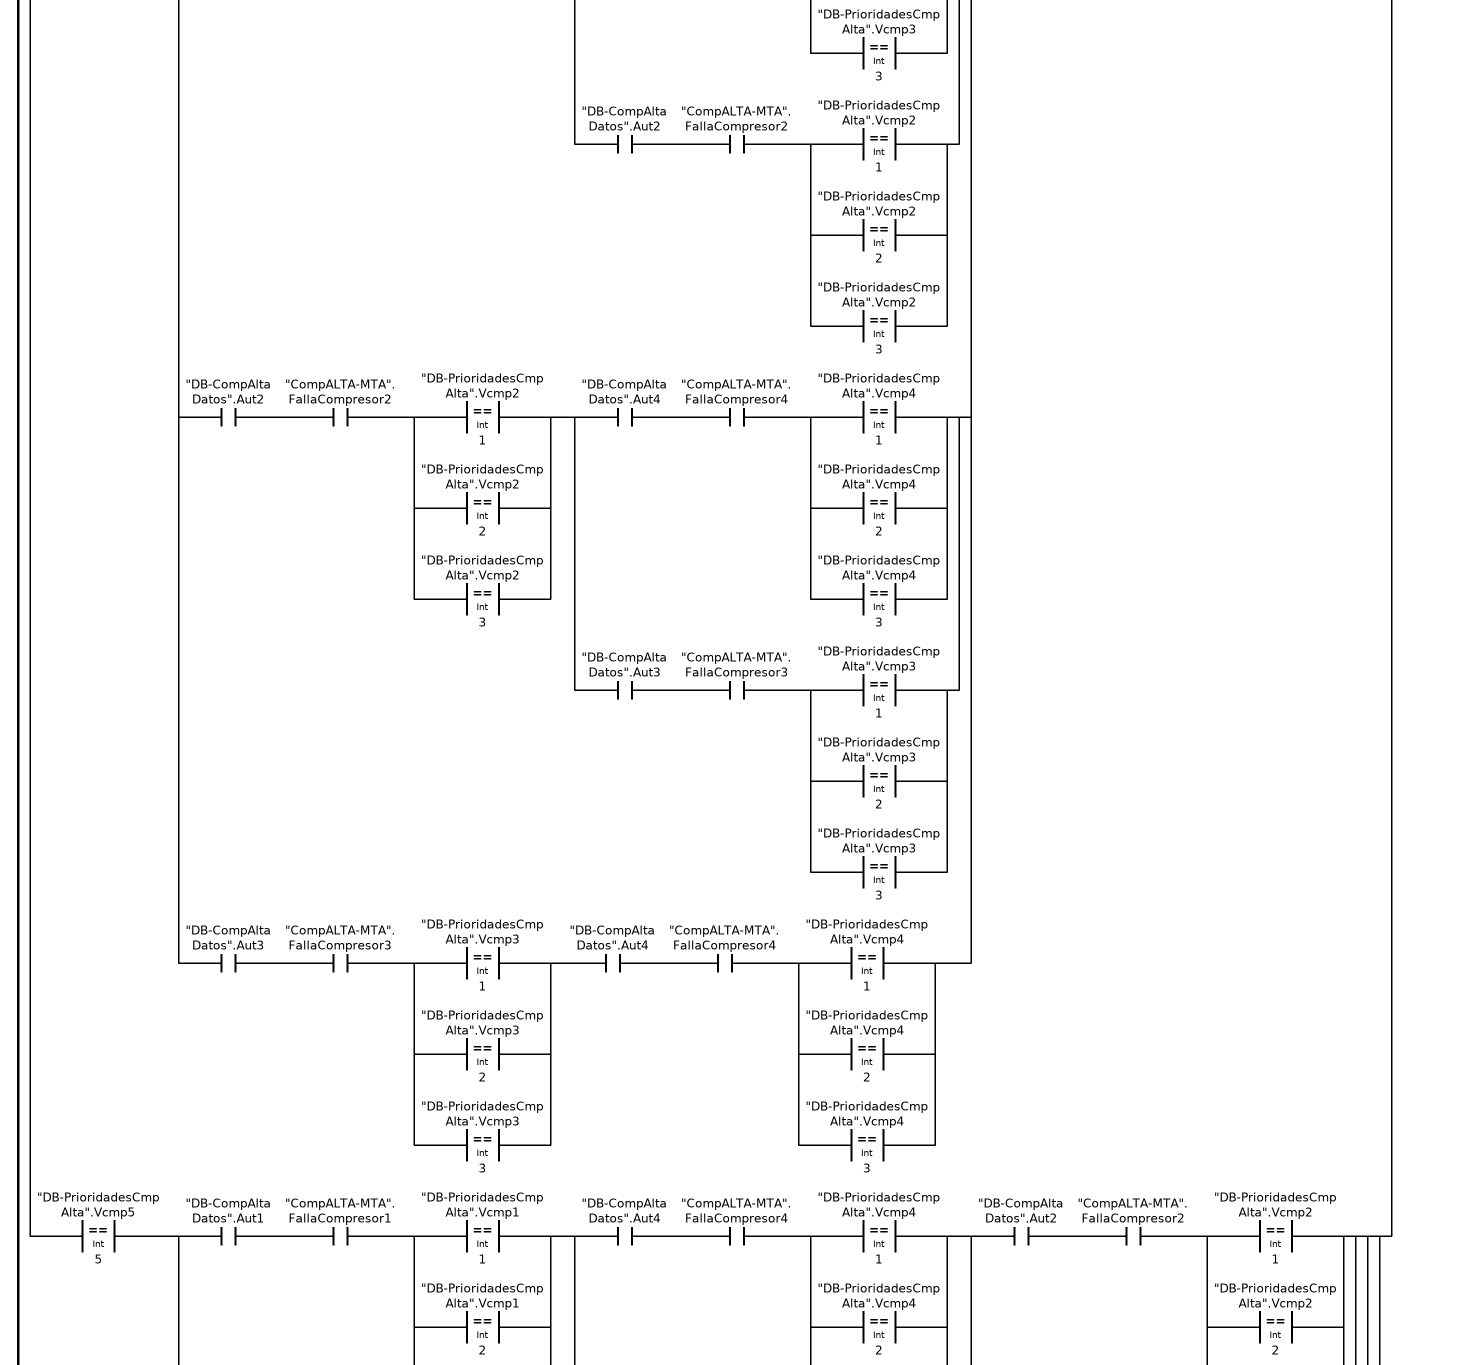
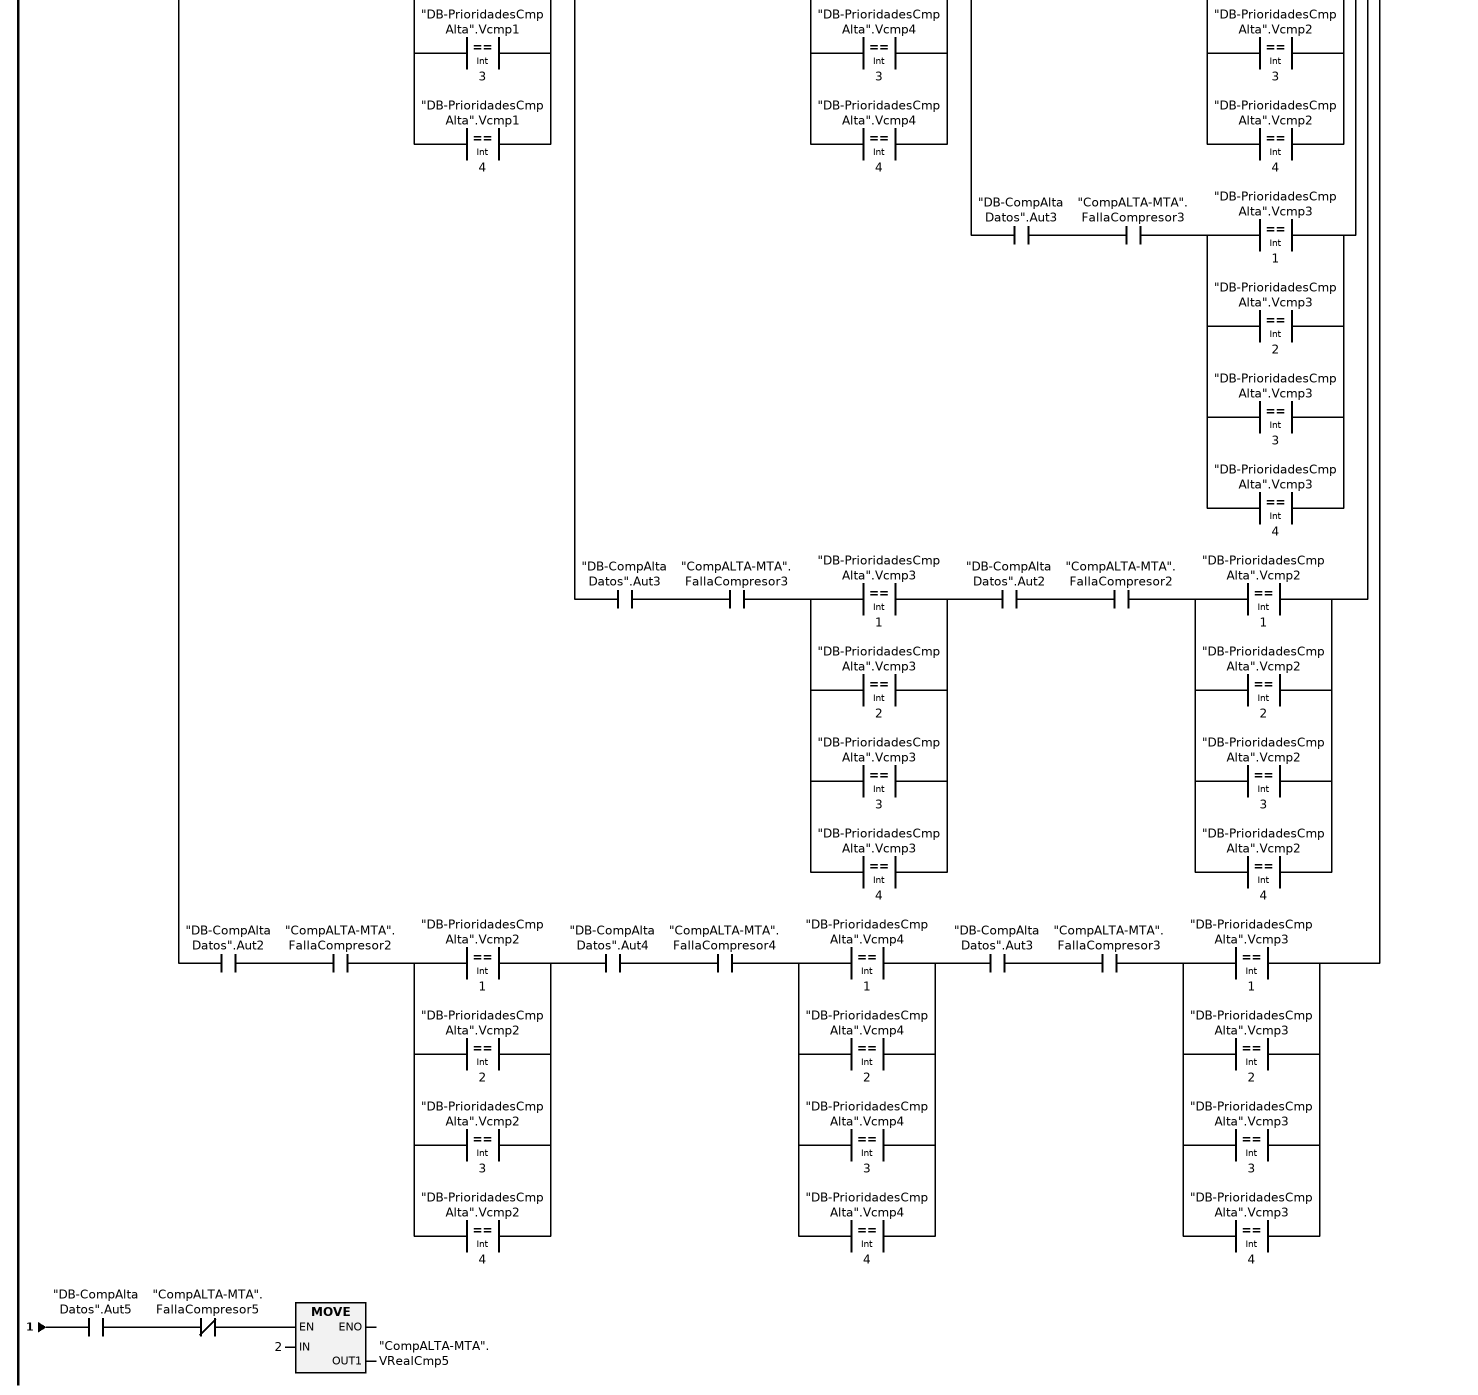
   IF (("DB-PrioridadesCmpAlta".Vcmp5 = 2) OR (("DB-PrioridadesCmpAlta".Vcmp5 = 3) AND (("DB-CompAltaDatos".Aut1 AND "CompALTA-MTA".FallaCompresor1 AND (("DB-PrioridadesCmpAlta".Vcmp1 = 2) OR ("DB-PrioridadesCmpAlta".Vcmp1 = 1))) OR ("DB-CompAltaDatos".Aut2 AND "CompALTA-MTA".FallaCompresor2 AND (("DB-PrioridadesCmpAlta".Vcmp2 = 2) OR ("DB-PrioridadesCmpAlta".Vcmp2 = 1))) OR ("DB-CompAltaDatos".Aut3 AND "CompALTA-MTA".FallaCompresor3 AND (("DB-PrioridadesCmpAlta".Vcmp3 = 2) OR ("DB-PrioridadesCmpAlta".Vcmp3 = 1))) OR ("DB-CompAltaDatos".Aut4 AND "CompALTA-MTA".FallaCompresor4 AND (("DB-PrioridadesCmpAlta".Vcmp4 = 2) OR ("DB-PrioridadesCmpAlta".Vcmp4 = 1))))) OR (("DB-PrioridadesCmpAlta".Vcmp5 = 4) AND (("DB-CompAltaDatos".Aut1 AND "CompALTA-MTA".FallaCompresor1 AND (("DB-PrioridadesCmpAlta".Vcmp1 = 1) OR ("DB-PrioridadesCmpAlta".Vcmp1 = 2) OR ("DB-PrioridadesCmpAlta".Vcmp1 = 3)) AND (("DB-CompAltaDatos".Aut4 AND "CompALTA-MTA".FallaCompresor4 AND (("DB-PrioridadesCmpAlta".Vcmp4 = 1) OR ("DB-PrioridadesCmpAlta".Vcmp4 = 2) OR ("DB-PrioridadesCmpAlta".Vcmp4 = 3))) OR ("DB-CompAltaDatos".Aut3 AND "CompALTA-MTA".FallaCompresor3 AND (("DB-PrioridadesCmpAlta".Vcmp3 = 1) OR ("DB-PrioridadesCmpAlta".Vcmp3 = 2) OR ("DB-PrioridadesCmpAlta".Vcmp3 = 3))) OR ("DB-CompAltaDatos".Aut2 AND "CompALTA-MTA".FallaCompresor2 AND (("DB-PrioridadesCmpAlta".Vcmp2 = 1) OR ("DB-PrioridadesCmpAlta".Vcmp2 = 2) OR ("DB-PrioridadesCmpAlta".Vcmp2 = 3))))) OR ("DB-CompAltaDatos".Aut2 AND "CompALTA-MTA".FallaCompresor2 AND (("DB-PrioridadesCmpAlta".Vcmp2 = 1) OR ("DB-PrioridadesCmpAlta".Vcmp2 = 2) OR ("DB-PrioridadesCmpAlta".Vcmp2 = 3)) AND (("DB-CompAltaDatos".Aut4 AND "CompALTA-MTA".FallaCompresor4 AND (("DB-PrioridadesCmpAlta".Vcmp4 = 1) OR ("DB-PrioridadesCmpAlta".Vcmp4 = 2) OR ("DB-PrioridadesCmpAlta".Vcmp4 = 3))) OR ("DB-CompAltaDatos".Aut3 AND "CompALTA-MTA".FallaCompresor3 AND (("DB-PrioridadesCmpAlta".Vcmp3 = 1) OR ("DB-PrioridadesCmpAlta".Vcmp3 = 2) OR ("DB-PrioridadesCmpAlta".Vcmp3 = 3))))) OR ("DB-CompAltaDatos".Aut3 AND "CompALTA-MTA".FallaCompresor3 AND (("DB-PrioridadesCmpAlta".Vcmp3 = 1) OR ("DB-PrioridadesCmpAlta".Vcmp3 = 2) OR ("DB-PrioridadesCmpAlta".Vcmp3 = 3)) AND "DB-CompAltaDatos".Aut4 AND "CompALTA-MTA".FallaCompresor4 AND (("DB-PrioridadesCmpAlta".Vcmp4 = 1) OR ("DB-PrioridadesCmpAlta".Vcmp4 = 2) OR ("DB-PrioridadesCmpAlta".Vcmp4 = 3))))) OR (("DB-PrioridadesCmpAlta".Vcmp5 = 5) AND (("DB-CompAltaDatos".Aut1 AND "CompALTA-MTA".FallaCompresor1 AND (("DB-PrioridadesCmpAlta".Vcmp1 = 1) OR ("DB-PrioridadesCmpAlta".Vcmp1 = 2) OR ("DB-PrioridadesCmpAlta".Vcmp1 = 3) OR ("DB-PrioridadesCmpAlta".Vcmp1 = 4)) AND (("DB-CompAltaDatos".Aut4 AND "CompALTA-MTA".FallaCompresor4 AND (("DB-PrioridadesCmpAlta".Vcmp4 = 1) OR ("DB-PrioridadesCmpAlta".Vcmp4 = 2) OR ("DB-PrioridadesCmpAlta".Vcmp4 = 3) OR ("DB-PrioridadesCmpAlta".Vcmp4 = 4)) AND (("DB-CompAltaDatos".Aut2 AND "CompALTA-MTA".FallaCompresor2 AND (("DB-PrioridadesCmpAlta".Vcmp2 = 1) OR ("DB-PrioridadesCmpAlta".Vcmp2 = 2) OR ("DB-PrioridadesCmpAlta".Vcmp2 = 3) OR ("DB-PrioridadesCmpAlta".Vcmp2 = 4))) OR ("DB-CompAltaDatos".Aut3 AND "CompALTA-MTA".FallaCompresor3 AND (("DB-PrioridadesCmpAlta".Vcmp3 = 1) OR ("DB-PrioridadesCmpAlta".Vcmp3 = 2) OR ("DB-PrioridadesCmpAlta".Vcmp3 = 3) OR ("DB-PrioridadesCmpAlta".Vcmp3 = 4))))) OR ("DB-CompAltaDatos".Aut3 AND "CompALTA-MTA".FallaCompresor3 AND (("DB-PrioridadesCmpAlta".Vcmp3 = 1) OR ("DB-PrioridadesCmpAlta".Vcmp3 = 2) OR ("DB-PrioridadesCmpAlta".Vcmp3 = 3) OR ("DB-PrioridadesCmpAlta".Vcmp3 = 4)) AND "DB-CompAltaDatos".Aut2 AND "CompALTA-MTA".FallaCompresor2 AND (("DB-PrioridadesCmpAlta".Vcmp2 = 1) OR ("DB-PrioridadesCmpAlta".Vcmp2 = 2) OR ("DB-PrioridadesCmpAlta".Vcmp2 = 3) OR ("DB-PrioridadesCmpAlta".Vcmp2 = 4))))) OR ("DB-CompAltaDatos".Aut2 AND "CompALTA-MTA".FallaCompresor2 AND (("DB-PrioridadesCmpAlta".Vcmp2 = 1) OR ("DB-PrioridadesCmpAlta".Vcmp2 = 2) OR ("DB-PrioridadesCmpAlta".Vcmp2 = 3) OR ("DB-PrioridadesCmpAlta".Vcmp2 = 4)) AND "DB-CompAltaDatos".Aut4 AND "CompALTA-MTA".FallaCompresor4 AND (("DB-PrioridadesCmpAlta".Vcmp4 = 1) OR ("DB-PrioridadesCmpAlta".Vcmp4 = 2) OR ("DB-PrioridadesCmpAlta".Vcmp4 = 3) OR ("DB-PrioridadesCmpAlta".Vcmp4 = 4)) AND "DB-CompAltaDatos".Aut3 AND "CompALTA-MTA".FallaCompresor3 AND (("DB-PrioridadesCmpAlta".Vcmp3 = 1) OR ("DB-PrioridadesCmpAlta".Vcmp3 = 2) OR ("DB-PrioridadesCmpAlta".Vcmp3 = 3) OR ("DB-PrioridadesCmpAlta".Vcmp3 = 4)))))) AND "DB-CompAltaDatos".Aut5 AND NOT "CompALTA-MTA".FallaCompresor5 THEN
       "CompALTA-MTA".VRealCmp5 := 2;
   END_IF;
END_REGION

REGION Network 33
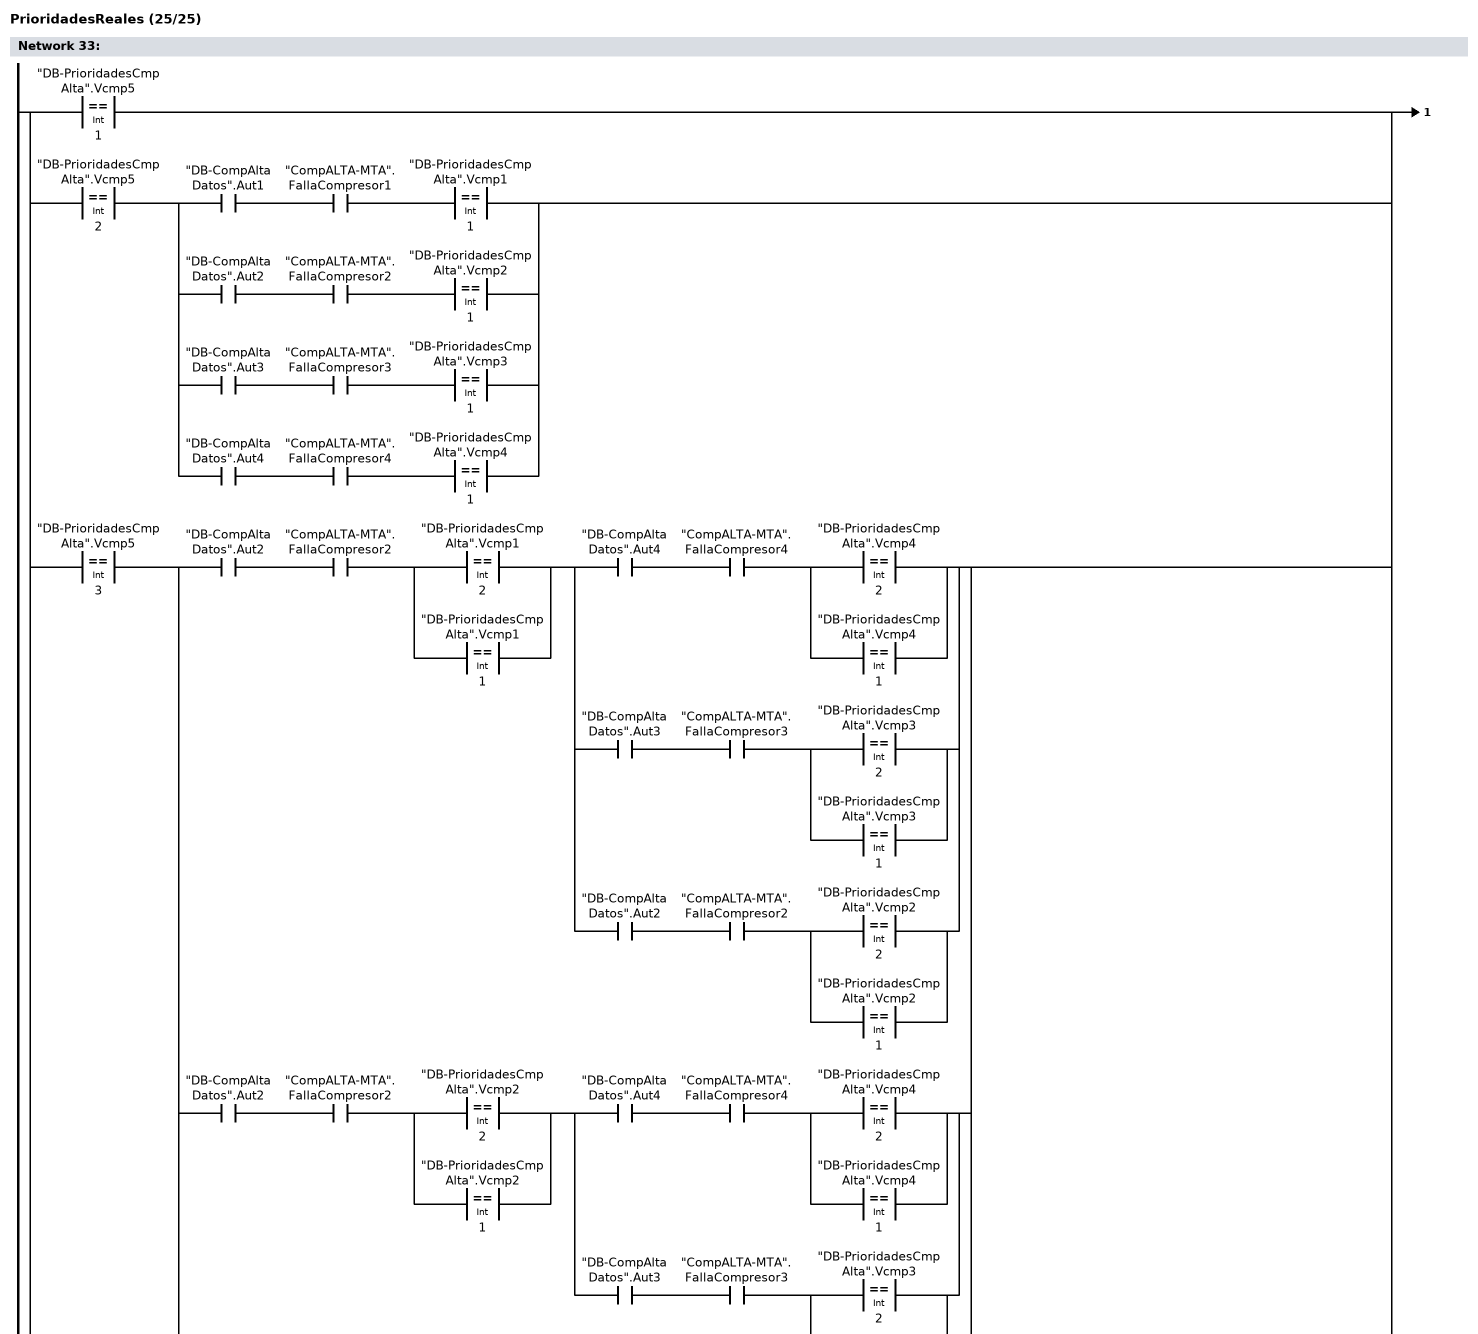
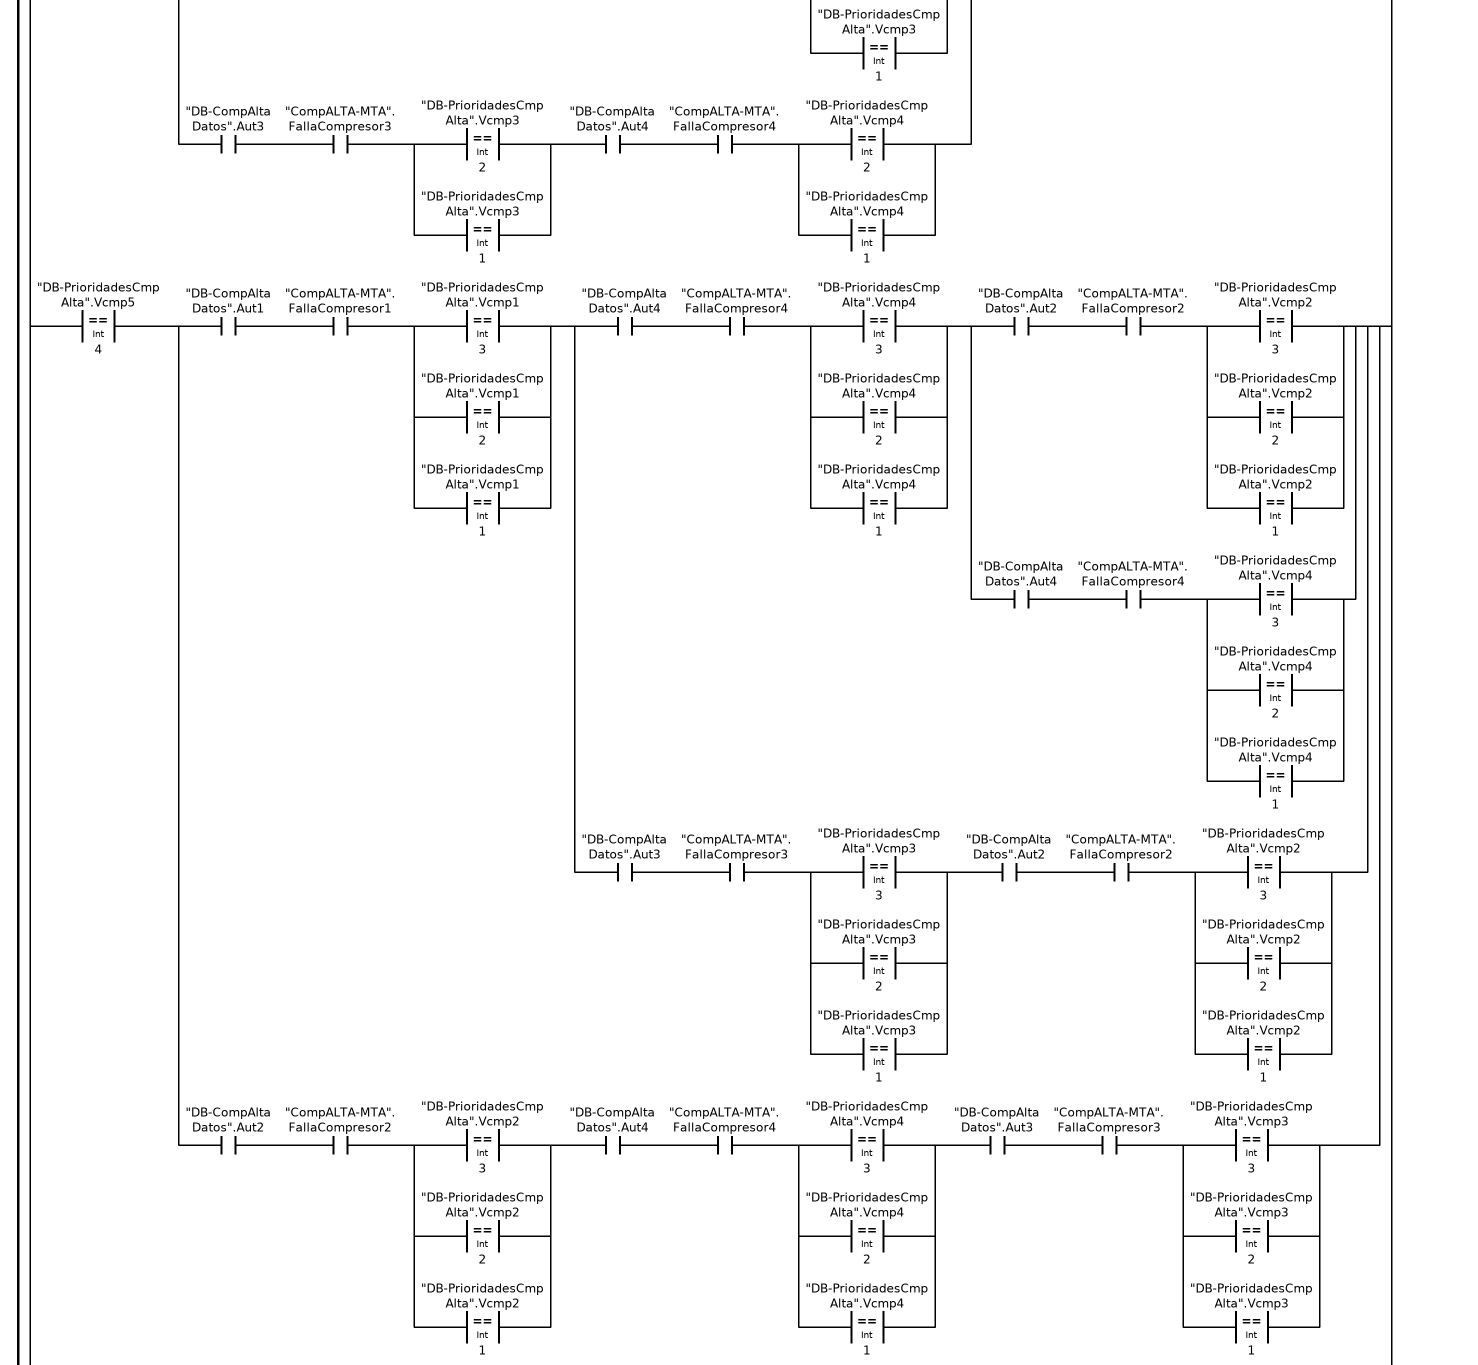
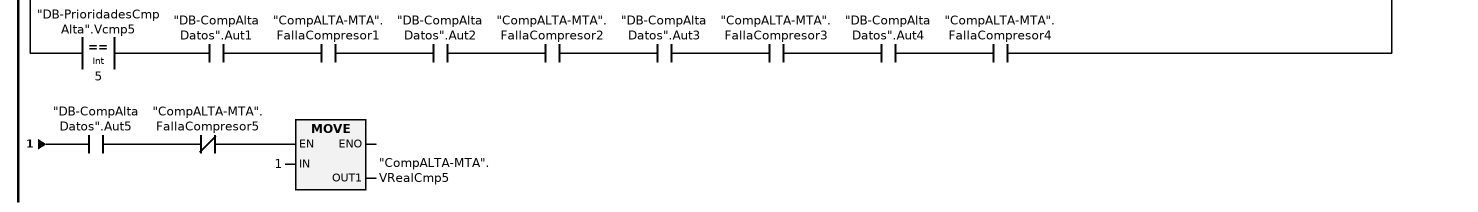
   IF (("DB-PrioridadesCmpAlta".Vcmp5 = 1) OR (("DB-PrioridadesCmpAlta".Vcmp5 = 2) AND (("DB-CompAltaDatos".Aut1 AND "CompALTA-MTA".FallaCompresor1 AND ("DB-PrioridadesCmpAlta".Vcmp1 = 1)) OR ("DB-CompAltaDatos".Aut2 AND "CompALTA-MTA".FallaCompresor2 AND ("DB-PrioridadesCmpAlta".Vcmp2 = 1)) OR ("DB-CompAltaDatos".Aut3 AND "CompALTA-MTA".FallaCompresor3 AND ("DB-PrioridadesCmpAlta".Vcmp3 = 1)) OR ("DB-CompAltaDatos".Aut4 AND "CompALTA-MTA".FallaCompresor4 AND ("DB-PrioridadesCmpAlta".Vcmp4 = 1)))) OR (("DB-PrioridadesCmpAlta".Vcmp5 = 3) AND (("DB-CompAltaDatos".Aut2 AND "CompALTA-MTA".FallaCompresor2 AND (("DB-PrioridadesCmpAlta".Vcmp1 = 2) OR ("DB-PrioridadesCmpAlta".Vcmp1 = 1)) AND (("DB-CompAltaDatos".Aut4 AND "CompALTA-MTA".FallaCompresor4 AND (("DB-PrioridadesCmpAlta".Vcmp4 = 2) OR ("DB-PrioridadesCmpAlta".Vcmp4 = 1))) OR ("DB-CompAltaDatos".Aut3 AND "CompALTA-MTA".FallaCompresor3 AND (("DB-PrioridadesCmpAlta".Vcmp3 = 2) OR ("DB-PrioridadesCmpAlta".Vcmp3 = 1))) OR ("DB-CompAltaDatos".Aut2 AND "CompALTA-MTA".FallaCompresor2 AND (("DB-PrioridadesCmpAlta".Vcmp2 = 2) OR ("DB-PrioridadesCmpAlta".Vcmp2 = 1))))) OR ("DB-CompAltaDatos".Aut2 AND "CompALTA-MTA".FallaCompresor2 AND (("DB-PrioridadesCmpAlta".Vcmp2 = 2) OR ("DB-PrioridadesCmpAlta".Vcmp2 = 1)) AND (("DB-CompAltaDatos".Aut4 AND "CompALTA-MTA".FallaCompresor4 AND (("DB-PrioridadesCmpAlta".Vcmp4 = 2) OR ("DB-PrioridadesCmpAlta".Vcmp4 = 1))) OR ("DB-CompAltaDatos".Aut3 AND "CompALTA-MTA".FallaCompresor3 AND (("DB-PrioridadesCmpAlta".Vcmp3 = 2) OR ("DB-PrioridadesCmpAlta".Vcmp3 = 1))))) OR ("DB-CompAltaDatos".Aut3 AND "CompALTA-MTA".FallaCompresor3 AND (("DB-PrioridadesCmpAlta".Vcmp3 = 2) OR ("DB-PrioridadesCmpAlta".Vcmp3 = 1)) AND "DB-CompAltaDatos".Aut4 AND "CompALTA-MTA".FallaCompresor4 AND (("DB-PrioridadesCmpAlta".Vcmp4 = 2) OR ("DB-PrioridadesCmpAlta".Vcmp4 = 1))))) OR (("DB-PrioridadesCmpAlta".Vcmp5 = 4) AND (("DB-CompAltaDatos".Aut1 AND "CompALTA-MTA".FallaCompresor1 AND (("DB-PrioridadesCmpAlta".Vcmp1 = 3) OR ("DB-PrioridadesCmpAlta".Vcmp1 = 2) OR ("DB-PrioridadesCmpAlta".Vcmp1 = 1)) AND (("DB-CompAltaDatos".Aut4 AND "CompALTA-MTA".FallaCompresor4 AND (("DB-PrioridadesCmpAlta".Vcmp4 = 3) OR ("DB-PrioridadesCmpAlta".Vcmp4 = 2) OR ("DB-PrioridadesCmpAlta".Vcmp4 = 1)) AND (("DB-CompAltaDatos".Aut2 AND "CompALTA-MTA".FallaCompresor2 AND (("DB-PrioridadesCmpAlta".Vcmp2 = 3) OR ("DB-PrioridadesCmpAlta".Vcmp2 = 2) OR ("DB-PrioridadesCmpAlta".Vcmp2 = 1))) OR ("DB-CompAltaDatos".Aut4 AND "CompALTA-MTA".FallaCompresor4 AND (("DB-PrioridadesCmpAlta".Vcmp4 = 3) OR ("DB-PrioridadesCmpAlta".Vcmp4 = 2) OR ("DB-PrioridadesCmpAlta".Vcmp4 = 1))))) OR ("DB-CompAltaDatos".Aut3 AND "CompALTA-MTA".FallaCompresor3 AND (("DB-PrioridadesCmpAlta".Vcmp3 = 3) OR ("DB-PrioridadesCmpAlta".Vcmp3 = 2) OR ("DB-PrioridadesCmpAlta".Vcmp3 = 1)) AND "DB-CompAltaDatos".Aut2 AND "CompALTA-MTA".FallaCompresor2 AND (("DB-PrioridadesCmpAlta".Vcmp2 = 3) OR ("DB-PrioridadesCmpAlta".Vcmp2 = 2) OR ("DB-PrioridadesCmpAlta".Vcmp2 = 1))))) OR ("DB-CompAltaDatos".Aut2 AND "CompALTA-MTA".FallaCompresor2 AND (("DB-PrioridadesCmpAlta".Vcmp2 = 3) OR ("DB-PrioridadesCmpAlta".Vcmp2 = 2) OR ("DB-PrioridadesCmpAlta".Vcmp2 = 1)) AND "DB-CompAltaDatos".Aut4 AND "CompALTA-MTA".FallaCompresor4 AND (("DB-PrioridadesCmpAlta".Vcmp4 = 3) OR ("DB-PrioridadesCmpAlta".Vcmp4 = 2) OR ("DB-PrioridadesCmpAlta".Vcmp4 = 1)) AND "DB-CompAltaDatos".Aut3 AND "CompALTA-MTA".FallaCompresor3 AND (("DB-PrioridadesCmpAlta".Vcmp3 = 3) OR ("DB-PrioridadesCmpAlta".Vcmp3 = 2) OR ("DB-PrioridadesCmpAlta".Vcmp3 = 1))))) OR (("DB-PrioridadesCmpAlta".Vcmp5 = 5) AND "DB-CompAltaDatos".Aut1 AND "CompALTA-MTA".FallaCompresor1 AND "DB-CompAltaDatos".Aut2 AND "CompALTA-MTA".FallaCompresor2 AND "DB-CompAltaDatos".Aut3 AND "CompALTA-MTA".FallaCompresor3 AND "DB-CompAltaDatos".Aut4 AND "CompALTA-MTA".FallaCompresor4)) AND "DB-CompAltaDatos".Aut5 AND NOT "CompALTA-MTA".FallaCompresor5 THEN
       "CompALTA-MTA".VRealCmp5 := 1;
   END_IF;
END_REGION
END_FUNCTION

FUNCTION "FlancosCmpAlta" : Void   // FC45, LAD
{ S7_Optimized_Access := 'FALSE' }
VERSION : 0.1
   VAR_TEMP   // added for the SCL form of the ladder/FBD networks
      _w1 : Bool;
      _w2 : Bool;
      _w3 : Bool;
      _w4 : Bool;
      _w5 : Bool;
      _w6 : Bool;
      _w7 : Bool;
      _s5time1 : S5Time;
   END_VAR
BEGIN

REGION Network 1
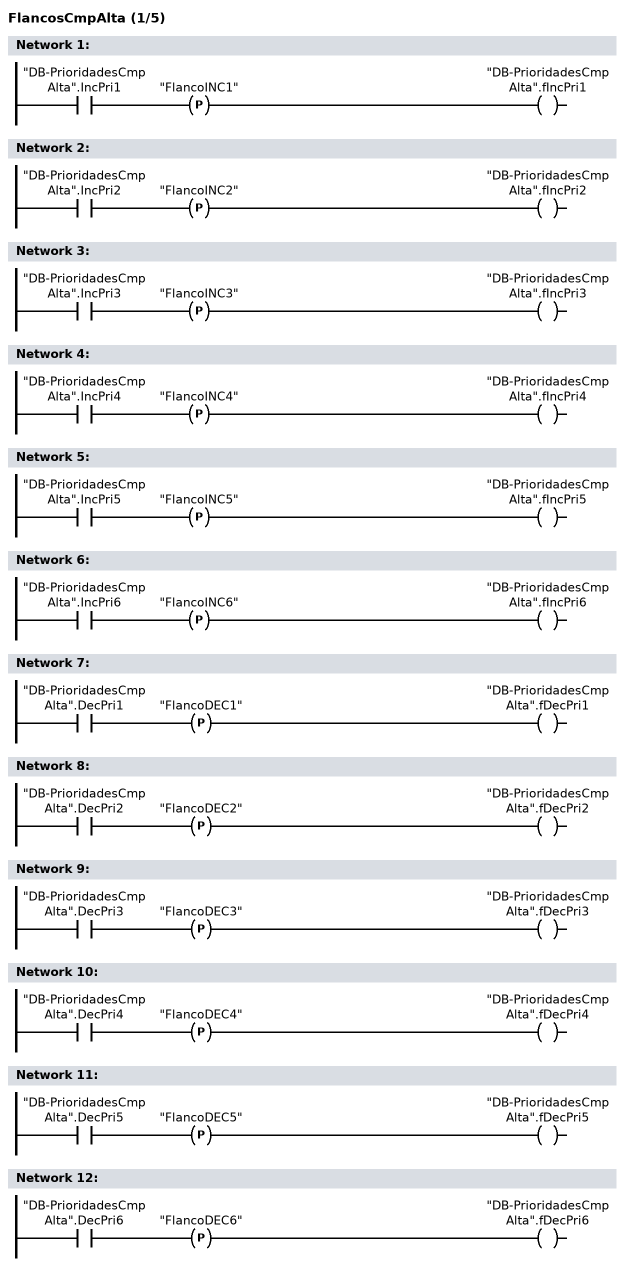
   RUNG wire#powerrail
      Contact( "DB-PrioridadesCmpAlta".IncPri1 )
      P_Trig( "FlancoINC1" )
      Coil( "DB-PrioridadesCmpAlta".fIncPri1 )
   END_RUNG
   // the same network as SCL:
   #_w1 := "DB-PrioridadesCmpAlta".IncPri1 AND NOT "FlancoINC1";   // rising edge
   "FlancoINC1" := "DB-PrioridadesCmpAlta".IncPri1;
   "DB-PrioridadesCmpAlta".fIncPri1 := #_w1;
END_REGION

REGION Network 2
   RUNG wire#powerrail
      Contact( "DB-PrioridadesCmpAlta".IncPri2 )
      P_Trig( "FlancoINC2" )
      Coil( "DB-PrioridadesCmpAlta".fIncPri2 )
   END_RUNG
   // the same network as SCL:
   #_w1 := "DB-PrioridadesCmpAlta".IncPri2 AND NOT "FlancoINC2";   // rising edge
   "FlancoINC2" := "DB-PrioridadesCmpAlta".IncPri2;
   "DB-PrioridadesCmpAlta".fIncPri2 := #_w1;
END_REGION

REGION Network 3
   RUNG wire#powerrail
      Contact( "DB-PrioridadesCmpAlta".IncPri3 )
      P_Trig( "FlancoINC3" )
      Coil( "DB-PrioridadesCmpAlta".fIncPri3 )
   END_RUNG
   // the same network as SCL:
   #_w1 := "DB-PrioridadesCmpAlta".IncPri3 AND NOT "FlancoINC3";   // rising edge
   "FlancoINC3" := "DB-PrioridadesCmpAlta".IncPri3;
   "DB-PrioridadesCmpAlta".fIncPri3 := #_w1;
END_REGION

REGION Network 4
   RUNG wire#powerrail
      Contact( "DB-PrioridadesCmpAlta".IncPri4 )
      P_Trig( "FlancoINC4" )
      Coil( "DB-PrioridadesCmpAlta".fIncPri4 )
   END_RUNG
   // the same network as SCL:
   #_w1 := "DB-PrioridadesCmpAlta".IncPri4 AND NOT "FlancoINC4";   // rising edge
   "FlancoINC4" := "DB-PrioridadesCmpAlta".IncPri4;
   "DB-PrioridadesCmpAlta".fIncPri4 := #_w1;
END_REGION

REGION Network 5
   RUNG wire#powerrail
      Contact( "DB-PrioridadesCmpAlta".IncPri5 )
      P_Trig( "FlancoINC5" )
      Coil( "DB-PrioridadesCmpAlta".fIncPri5 )
   END_RUNG
   // the same network as SCL:
   #_w1 := "DB-PrioridadesCmpAlta".IncPri5 AND NOT "FlancoINC5";   // rising edge
   "FlancoINC5" := "DB-PrioridadesCmpAlta".IncPri5;
   "DB-PrioridadesCmpAlta".fIncPri5 := #_w1;
END_REGION

REGION Network 6
   RUNG wire#powerrail
      Contact( "DB-PrioridadesCmpAlta".IncPri6 )
      P_Trig( "FlancoINC6" )
      Coil( "DB-PrioridadesCmpAlta".fIncPri6 )
   END_RUNG
   // the same network as SCL:
   #_w1 := "DB-PrioridadesCmpAlta".IncPri6 AND NOT "FlancoINC6";   // rising edge
   "FlancoINC6" := "DB-PrioridadesCmpAlta".IncPri6;
   "DB-PrioridadesCmpAlta".fIncPri6 := #_w1;
END_REGION

REGION Network 7
   RUNG wire#powerrail
      Contact( "DB-PrioridadesCmpAlta".DecPri1 )
      P_Trig( "FlancoDEC1" )
      Coil( "DB-PrioridadesCmpAlta".fDecPri1 )
   END_RUNG
   // the same network as SCL:
   #_w1 := "DB-PrioridadesCmpAlta".DecPri1 AND NOT "FlancoDEC1";   // rising edge
   "FlancoDEC1" := "DB-PrioridadesCmpAlta".DecPri1;
   "DB-PrioridadesCmpAlta".fDecPri1 := #_w1;
END_REGION

REGION Network 8
   RUNG wire#powerrail
      Contact( "DB-PrioridadesCmpAlta".DecPri2 )
      P_Trig( "FlancoDEC2" )
      Coil( "DB-PrioridadesCmpAlta".fDecPri2 )
   END_RUNG
   // the same network as SCL:
   #_w1 := "DB-PrioridadesCmpAlta".DecPri2 AND NOT "FlancoDEC2";   // rising edge
   "FlancoDEC2" := "DB-PrioridadesCmpAlta".DecPri2;
   "DB-PrioridadesCmpAlta".fDecPri2 := #_w1;
END_REGION

REGION Network 9
   RUNG wire#powerrail
      Contact( "DB-PrioridadesCmpAlta".DecPri3 )
      P_Trig( "FlancoDEC3" )
      Coil( "DB-PrioridadesCmpAlta".fDecPri3 )
   END_RUNG
   // the same network as SCL:
   #_w1 := "DB-PrioridadesCmpAlta".DecPri3 AND NOT "FlancoDEC3";   // rising edge
   "FlancoDEC3" := "DB-PrioridadesCmpAlta".DecPri3;
   "DB-PrioridadesCmpAlta".fDecPri3 := #_w1;
END_REGION

REGION Network 10
   RUNG wire#powerrail
      Contact( "DB-PrioridadesCmpAlta".DecPri4 )
      P_Trig( "FlancoDEC4" )
      Coil( "DB-PrioridadesCmpAlta".fDecPri4 )
   END_RUNG
   // the same network as SCL:
   #_w1 := "DB-PrioridadesCmpAlta".DecPri4 AND NOT "FlancoDEC4";   // rising edge
   "FlancoDEC4" := "DB-PrioridadesCmpAlta".DecPri4;
   "DB-PrioridadesCmpAlta".fDecPri4 := #_w1;
END_REGION

REGION Network 11
   RUNG wire#powerrail
      Contact( "DB-PrioridadesCmpAlta".DecPri5 )
      P_Trig( "FlancoDEC5" )
      Coil( "DB-PrioridadesCmpAlta".fDecPri5 )
   END_RUNG
   // the same network as SCL:
   #_w1 := "DB-PrioridadesCmpAlta".DecPri5 AND NOT "FlancoDEC5";   // rising edge
   "FlancoDEC5" := "DB-PrioridadesCmpAlta".DecPri5;
   "DB-PrioridadesCmpAlta".fDecPri5 := #_w1;
END_REGION

REGION Network 12
   RUNG wire#powerrail
      Contact( "DB-PrioridadesCmpAlta".DecPri6 )
      P_Trig( "FlancoDEC6" )
      Coil( "DB-PrioridadesCmpAlta".fDecPri6 )
   END_RUNG
   // the same network as SCL:
   #_w1 := "DB-PrioridadesCmpAlta".DecPri6 AND NOT "FlancoDEC6";   // rising edge
   "FlancoDEC6" := "DB-PrioridadesCmpAlta".DecPri6;
   "DB-PrioridadesCmpAlta".fDecPri6 := #_w1;
END_REGION

REGION Network 13
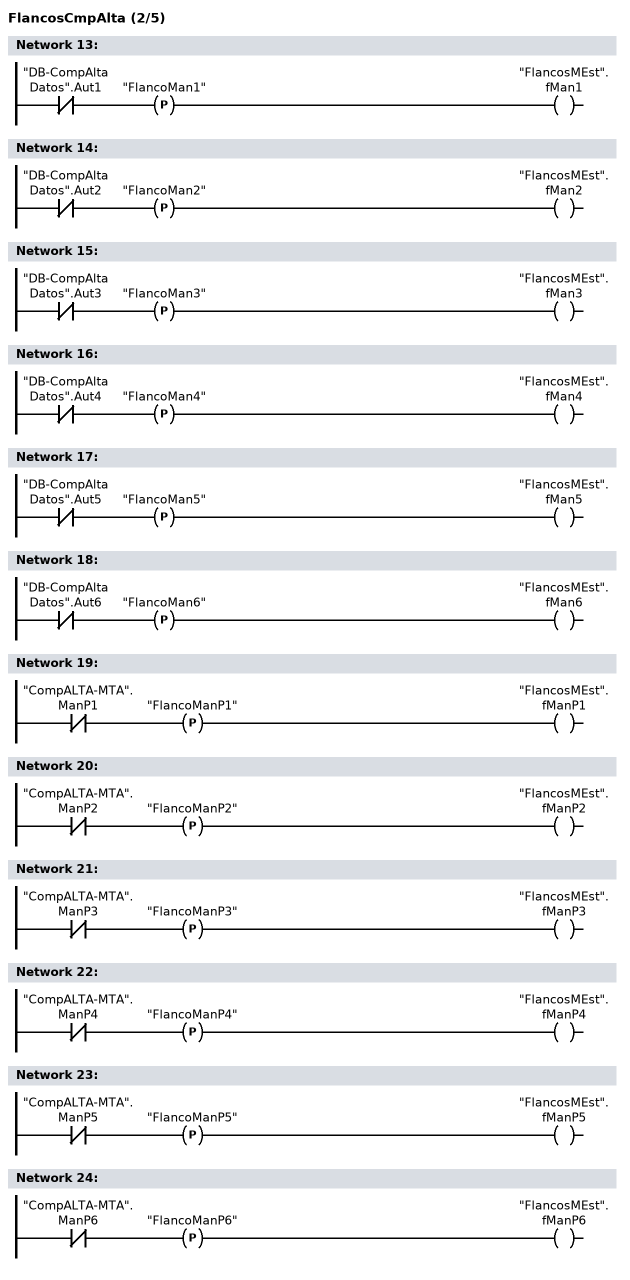
   RUNG wire#powerrail
      I_Contact( "DB-CompAltaDatos".Aut1 )
      P_Trig( "FlancoMan1" )
      Coil( "FlancosMEst".fMan1 )
   END_RUNG
   // the same network as SCL:
   #_w1 := NOT "DB-CompAltaDatos".Aut1 AND NOT "FlancoMan1";   // rising edge
   "FlancoMan1" := NOT "DB-CompAltaDatos".Aut1;
   "FlancosMEst".fMan1 := #_w1;
END_REGION

REGION Network 14
   RUNG wire#powerrail
      I_Contact( "DB-CompAltaDatos".Aut2 )
      P_Trig( "FlancoMan2" )
      Coil( "FlancosMEst".fMan2 )
   END_RUNG
   // the same network as SCL:
   #_w1 := NOT "DB-CompAltaDatos".Aut2 AND NOT "FlancoMan2";   // rising edge
   "FlancoMan2" := NOT "DB-CompAltaDatos".Aut2;
   "FlancosMEst".fMan2 := #_w1;
END_REGION

REGION Network 15
   RUNG wire#powerrail
      I_Contact( "DB-CompAltaDatos".Aut3 )
      P_Trig( "FlancoMan3" )
      Coil( "FlancosMEst".fMan3 )
   END_RUNG
   // the same network as SCL:
   #_w1 := NOT "DB-CompAltaDatos".Aut3 AND NOT "FlancoMan3";   // rising edge
   "FlancoMan3" := NOT "DB-CompAltaDatos".Aut3;
   "FlancosMEst".fMan3 := #_w1;
END_REGION

REGION Network 16
   RUNG wire#powerrail
      I_Contact( "DB-CompAltaDatos".Aut4 )
      P_Trig( "FlancoMan4" )
      Coil( "FlancosMEst".fMan4 )
   END_RUNG
   // the same network as SCL:
   #_w1 := NOT "DB-CompAltaDatos".Aut4 AND NOT "FlancoMan4";   // rising edge
   "FlancoMan4" := NOT "DB-CompAltaDatos".Aut4;
   "FlancosMEst".fMan4 := #_w1;
END_REGION

REGION Network 17
   RUNG wire#powerrail
      I_Contact( "DB-CompAltaDatos".Aut5 )
      P_Trig( "FlancoMan5" )
      Coil( "FlancosMEst".fMan5 )
   END_RUNG
   // the same network as SCL:
   #_w1 := NOT "DB-CompAltaDatos".Aut5 AND NOT "FlancoMan5";   // rising edge
   "FlancoMan5" := NOT "DB-CompAltaDatos".Aut5;
   "FlancosMEst".fMan5 := #_w1;
END_REGION

REGION Network 18
   RUNG wire#powerrail
      I_Contact( "DB-CompAltaDatos".Aut6 )
      P_Trig( "FlancoMan6" )
      Coil( "FlancosMEst".fMan6 )
   END_RUNG
   // the same network as SCL:
   #_w1 := NOT "DB-CompAltaDatos".Aut6 AND NOT "FlancoMan6";   // rising edge
   "FlancoMan6" := NOT "DB-CompAltaDatos".Aut6;
   "FlancosMEst".fMan6 := #_w1;
END_REGION

REGION Network 19
   RUNG wire#powerrail
      I_Contact( "CompALTA-MTA".ManP1 )
      P_Trig( "FlancoManP1" )
      Coil( "FlancosMEst".fManP1 )
   END_RUNG
   // the same network as SCL:
   #_w1 := NOT "CompALTA-MTA".ManP1 AND NOT "FlancoManP1";   // rising edge
   "FlancoManP1" := NOT "CompALTA-MTA".ManP1;
   "FlancosMEst".fManP1 := #_w1;
END_REGION

REGION Network 20
   RUNG wire#powerrail
      I_Contact( "CompALTA-MTA".ManP2 )
      P_Trig( "FlancoManP2" )
      Coil( "FlancosMEst".fManP2 )
   END_RUNG
   // the same network as SCL:
   #_w1 := NOT "CompALTA-MTA".ManP2 AND NOT "FlancoManP2";   // rising edge
   "FlancoManP2" := NOT "CompALTA-MTA".ManP2;
   "FlancosMEst".fManP2 := #_w1;
END_REGION

REGION Network 21
   RUNG wire#powerrail
      I_Contact( "CompALTA-MTA".ManP3 )
      P_Trig( "FlancoManP3" )
      Coil( "FlancosMEst".fManP3 )
   END_RUNG
   // the same network as SCL:
   #_w1 := NOT "CompALTA-MTA".ManP3 AND NOT "FlancoManP3";   // rising edge
   "FlancoManP3" := NOT "CompALTA-MTA".ManP3;
   "FlancosMEst".fManP3 := #_w1;
END_REGION

REGION Network 22
   RUNG wire#powerrail
      I_Contact( "CompALTA-MTA".ManP4 )
      P_Trig( "FlancoManP4" )
      Coil( "FlancosMEst".fManP4 )
   END_RUNG
   // the same network as SCL:
   #_w1 := NOT "CompALTA-MTA".ManP4 AND NOT "FlancoManP4";   // rising edge
   "FlancoManP4" := NOT "CompALTA-MTA".ManP4;
   "FlancosMEst".fManP4 := #_w1;
END_REGION

REGION Network 23
   RUNG wire#powerrail
      I_Contact( "CompALTA-MTA".ManP5 )
      P_Trig( "FlancoManP5" )
      Coil( "FlancosMEst".fManP5 )
   END_RUNG
   // the same network as SCL:
   #_w1 := NOT "CompALTA-MTA".ManP5 AND NOT "FlancoManP5";   // rising edge
   "FlancoManP5" := NOT "CompALTA-MTA".ManP5;
   "FlancosMEst".fManP5 := #_w1;
END_REGION

REGION Network 24
   RUNG wire#powerrail
      I_Contact( "CompALTA-MTA".ManP6 )
      P_Trig( "FlancoManP6" )
      Coil( "FlancosMEst".fManP6 )
   END_RUNG
   // the same network as SCL:
   #_w1 := NOT "CompALTA-MTA".ManP6 AND NOT "FlancoManP6";   // rising edge
   "FlancoManP6" := NOT "CompALTA-MTA".ManP6;
   "FlancosMEst".fManP6 := #_w1;
END_REGION

REGION Network 25